      { S7_GenerateENO := "TRUE" } Add(in1 := "Archiwizowane_parametry".Wilgotnosc_srednia[0], in2 := "Archiwizowane_parametry".Wilgotnosc["Archiwizowane_parametry".iterator_srednia], out => "Archiwizowane_parametry".Wilgotnosc_srednia[0])
      Div(in1 := "Archiwizowane_parametry".Naslonecznienie_suma[0], in2 := "Archiwizowane_parametry".dzielnik, out => "Archiwizowane_parametry".Naslonecznienie_srednia[0])
      Div(in1 := "Archiwizowane_parametry".Temperatura_suma[0], in2 := "Archiwizowane_parametry".dzielnik, out => "Archiwizowane_parametry".Temperatura_srednia[0])
      Div(in1 := "Archiwizowane_parametry".Wilgotnosc_suma[0], in2 := "Archiwizowane_parametry".dzielnik, out => "Archiwizowane_parametry".Wilgotnosc_srednia[0])
   END_RUNG
   RUNG wire#w2
      { S7_Templates := "SrcType := Int" } GE_Contact(in1 := "Archiwizowane_parametry".iterator_srednia, in2 := 16)
      { S7_Templates := "SrcType := Int" } LT_Contact(in1 := "Archiwizowane_parametry".iterator_srednia, in2 := 32)
      { S7_GenerateENO := "TRUE" } Add(in1 := "Archiwizowane_parametry".Naslonecznienie_srednia[1], in2 := "Archiwizowane_parametry".Naslonecznienie["Archiwizowane_parametry".iterator_srednia], out => "Archiwizowane_parametry".Naslonecznienie_srednia[1])
      { S7_GenerateENO := "TRUE" } Add(in1 := "Archiwizowane_parametry".Temperatura_srednia[1], in2 := "Archiwizowane_parametry".Temperatura["Archiwizowane_parametry".iterator_srednia], out => "Archiwizowane_parametry".Temperatura_srednia[1])
      { S7_GenerateENO := "TRUE" } Add(in1 := "Archiwizowane_parametry".Wilgotnosc_srednia[1], in2 := "Archiwizowane_parametry".Wilgotnosc["Archiwizowane_parametry".iterator_srednia], out => "Archiwizowane_parametry".Wilgotnosc_srednia[1])
      Div(in1 := "Archiwizowane_parametry".Naslonecznienie_suma[1], in2 := "Archiwizowane_parametry".dzielnik, out => "Archiwizowane_parametry".Naslonecznienie_srednia[1])
      Div(in1 := "Archiwizowane_parametry".Temperatura_suma[1], in2 := "Archiwizowane_parametry".dzielnik, out => "Archiwizowane_parametry".Temperatura_srednia[1])
      Div(in1 := "Archiwizowane_parametry".Wilgotnosc_suma[1], in2 := "Archiwizowane_parametry".dzielnik, out => "Archiwizowane_parametry".Wilgotnosc_srednia[1])
   END_RUNG
   RUNG wire#w2
      { S7_Templates := "SrcType := Int" } GE_Contact(in1 := "Archiwizowane_parametry".iterator_srednia, in2 := 32)
      { S7_Templates := "SrcType := Int" } LT_Contact(in1 := "Archiwizowane_parametry".iterator_srednia, in2 := 48)
      { S7_GenerateENO := "TRUE" } Add(in1 := "Archiwizowane_parametry".Naslonecznienie_srednia[2], in2 := "Archiwizowane_parametry".Naslonecznienie["Archiwizowane_parametry".iterator_srednia], out => "Archiwizowane_parametry".Naslonecznienie_srednia[2])
      { S7_GenerateENO := "TRUE" } Add(in1 := "Archiwizowane_parametry".Temperatura_srednia[2], in2 := "Archiwizowane_parametry".Temperatura["Archiwizowane_parametry".iterator_srednia], out => "Archiwizowane_parametry".Temperatura_srednia[2])
      { S7_GenerateENO := "TRUE" } Add(in1 := "Archiwizowane_parametry".Wilgotnosc_srednia[2], in2 := "Archiwizowane_parametry".Wilgotnosc["Archiwizowane_parametry".iterator_srednia], out => "Archiwizowane_parametry".Wilgotnosc_srednia[2])
      Div(in1 := "Archiwizowane_parametry".Naslonecznienie_suma[2], in2 := "Archiwizowane_parametry".dzielnik, out => "Archiwizowane_parametry".Naslonecznienie_srednia[2])
      Div(in1 := "Archiwizowane_parametry".Temperatura_suma[2], in2 := "Archiwizowane_parametry".dzielnik, out => "Archiwizowane_parametry".Temperatura_srednia[2])
      Div(in1 := "Archiwizowane_parametry".Wilgotnosc_suma[2], in2 := "Archiwizowane_parametry".dzielnik, out => "Archiwizowane_parametry".Wilgotnosc_srednia[2])
   END_RUNG
   RUNG wire#w2
      { S7_Templates := "SrcType := Int" } GE_Contact(in1 := "Archiwizowane_parametry".iterator_srednia, in2 := 48)
      { S7_Templates := "SrcType := Int" } LT_Contact(in1 := "Archiwizowane_parametry".iterator_srednia, in2 := 64)
      { S7_GenerateENO := "TRUE" } Add(in1 := "Archiwizowane_parametry".Naslonecznienie_srednia[3], in2 := "Archiwizowane_parametry".Naslonecznienie["Archiwizowane_parametry".iterator_srednia], out => "Archiwizowane_parametry".Naslonecznienie_srednia[3])
      { S7_GenerateENO := "TRUE" } Add(in1 := "Archiwizowane_parametry".Temperatura_srednia[3], in2 := "Archiwizowane_parametry".Temperatura["Archiwizowane_parametry".iterator_srednia], out => "Archiwizowane_parametry".Temperatura_srednia[3])
      { S7_GenerateENO := "TRUE" } Add(in1 := "Archiwizowane_parametry".Wilgotnosc_srednia[3], in2 := "Archiwizowane_parametry".Wilgotnosc["Archiwizowane_parametry".iterator_srednia], out => "Archiwizowane_parametry".Wilgotnosc_srednia[3])
      Div(in1 := "Archiwizowane_parametry".Naslonecznienie_suma[3], in2 := "Archiwizowane_parametry".dzielnik, out => "Archiwizowane_parametry".Naslonecznienie_srednia[3])
      Div(in1 := "Archiwizowane_parametry".Temperatura_suma[3], in2 := "Archiwizowane_parametry".dzielnik, out => "Archiwizowane_parametry".Temperatura_srednia[3])
      Div(in1 := "Archiwizowane_parametry".Wilgotnosc_suma[3], in2 := "Archiwizowane_parametry".dzielnik, out => "Archiwizowane_parametry".Wilgotnosc_srednia[3])
   END_RUNG
   RUNG wire#w2
      { S7_Templates := "SrcType := Int" } GE_Contact(in1 := "Archiwizowane_parametry".iterator_srednia, in2 := 64)
      { S7_Templates := "SrcType := Int" } LT_Contact(in1 := "Archiwizowane_parametry".iterator_srednia, in2 := 80)
      { S7_GenerateENO := "TRUE" } Add(in1 := "Archiwizowane_parametry".Naslonecznienie_srednia[4], in2 := "Archiwizowane_parametry".Naslonecznienie["Archiwizowane_parametry".iterator_srednia], out => "Archiwizowane_parametry".Naslonecznienie_srednia[4])
      { S7_GenerateENO := "TRUE" } Add(in1 := "Archiwizowane_parametry".Temperatura_srednia[4], in2 := "Archiwizowane_parametry".Temperatura["Archiwizowane_parametry".iterator_srednia], out => "Archiwizowane_parametry".Temperatura_srednia[4])
      { S7_GenerateENO := "TRUE" } Add(in1 := "Archiwizowane_parametry".Wilgotnosc_srednia[4], in2 := "Archiwizowane_parametry".Wilgotnosc["Archiwizowane_parametry".iterator_srednia], out => "Archiwizowane_parametry".Wilgotnosc_srednia[4])
      Div(in1 := "Archiwizowane_parametry".Naslonecznienie_suma[4], in2 := "Archiwizowane_parametry".dzielnik, out => "Archiwizowane_parametry".Naslonecznienie_srednia[4])
      Div(in1 := "Archiwizowane_parametry".Temperatura_suma[4], in2 := "Archiwizowane_parametry".dzielnik, out => "Archiwizowane_parametry".Temperatura_srednia[4])
      Div(in1 := "Archiwizowane_parametry".Wilgotnosc_suma[4], in2 := "Archiwizowane_parametry".dzielnik, out => "Archiwizowane_parametry".Wilgotnosc_srednia[4])
   END_RUNG
   RUNG wire#w2
      { S7_Templates := "SrcType := Int" } GE_Contact(in1 := "Archiwizowane_parametry".iterator_srednia, in2 := 80)
      { S7_Templates := "SrcType := Int" } LT_Contact(in1 := "Archiwizowane_parametry".iterator_srednia, in2 := 96)
      { S7_GenerateENO := "TRUE" } Add(in1 := "Archiwizowane_parametry".Naslonecznienie_srednia[5], in2 := "Archiwizowane_parametry".Naslonecznienie["Archiwizowane_parametry".iterator_srednia], out => "Archiwizowane_parametry".Naslonecznienie_srednia[5])
      { S7_GenerateENO := "TRUE" } Add(in1 := "Archiwizowane_parametry".Temperatura_srednia[5], in2 := "Archiwizowane_parametry".Temperatura["Archiwizowane_parametry".iterator_srednia], out => "Archiwizowane_parametry".Temperatura_srednia[5])
      { S7_GenerateENO := "TRUE" } Add(in1 := "Archiwizowane_parametry".Wilgotnosc_srednia[5], in2 := "Archiwizowane_parametry".Wilgotnosc["Archiwizowane_parametry".iterator_srednia], out => "Archiwizowane_parametry".Wilgotnosc_srednia[5])
      Div(in1 := "Archiwizowane_parametry".Naslonecznienie_suma[5], in2 := "Archiwizowane_parametry".dzielnik, out => "Archiwizowane_parametry".Naslonecznienie_srednia[5])
      Div(in1 := "Archiwizowane_parametry".Temperatura_suma[5], in2 := "Archiwizowane_parametry".dzielnik, out => "Archiwizowane_parametry".Temperatura_srednia[5])
      Div(in1 := "Archiwizowane_parametry".Wilgotnosc_suma[5], in2 := "Archiwizowane_parametry".dzielnik, out => "Archiwizowane_parametry".Wilgotnosc_srednia[5])
   END_RUNG
   RUNG wire#w2
      { S7_Templates := "SrcType := Int" } GE_Contact(in1 := "Archiwizowane_parametry".iterator_srednia, in2 := 96)
      { S7_GenerateENO := "TRUE" } Add(in1 := "Archiwizowane_parametry".Naslonecznienie_srednia[6], in2 := "Archiwizowane_parametry".Naslonecznienie["Archiwizowane_parametry".iterator_srednia], out => "Archiwizowane_parametry".Naslonecznienie_srednia[6])
      { S7_GenerateENO := "TRUE" } Add(in1 := "Archiwizowane_parametry".Temperatura_srednia[6], in2 := "Archiwizowane_parametry".Temperatura["Archiwizowane_parametry".iterator_srednia], out => "Archiwizowane_parametry".Temperatura_srednia[6])
      { S7_GenerateENO := "TRUE" } Add(in1 := "Archiwizowane_parametry".Wilgotnosc_srednia[6], in2 := "Archiwizowane_parametry".Wilgotnosc["Archiwizowane_parametry".iterator_srednia], out => "Archiwizowane_parametry".Wilgotnosc_srednia[6])
      Div(in1 := "Archiwizowane_parametry".Naslonecznienie_suma[6], in2 := "Archiwizowane_parametry".dzielnik, out => "Archiwizowane_parametry".Naslonecznienie_srednia[6])
      Div(in1 := "Archiwizowane_parametry".Temperatura_suma[6], in2 := "Archiwizowane_parametry".dzielnik, out => "Archiwizowane_parametry".Temperatura_srednia[6])
      Div(in1 := "Archiwizowane_parametry".Wilgotnosc_suma[6], in2 := "Archiwizowane_parametry".dzielnik, out => "Archiwizowane_parametry".Wilgotnosc_srednia[6])
   END_RUNG
   RUNG wire#w1
      { S7_GenerateENO := "TRUE" } Add(in1 := "Archiwizowane_parametry".iterator_srednia, in2 := 1, out => "Archiwizowane_parametry".iterator_srednia)
   END_RUNG
   // the same network as SCL:
   // ENO of a box is taken as its EN; it also drops when the box reports an error
   #_w1 := "Archiwizowane_parametry".iterator_srednia < 112;
   #_w2 := #_w1 AND ("Archiwizowane_parametry".Wilgotnosc["Archiwizowane_parametry".iterator_srednia] >= 0);
   IF #_w2 THEN "Archiwizowane_parametry".dzielnik := "Archiwizowane_parametry".dzielnik + 1; END_IF;
   IF #_w2 AND ("Archiwizowane_parametry".iterator_srednia < 16) THEN
       "Archiwizowane_parametry".Naslonecznienie_srednia[0] := "Archiwizowane_parametry".Naslonecznienie_srednia[0] + "Archiwizowane_parametry".Naslonecznienie["Archiwizowane_parametry".iterator_srednia];
       "Archiwizowane_parametry".Temperatura_srednia[0] := "Archiwizowane_parametry".Temperatura_srednia[0] + "Archiwizowane_parametry".Temperatura["Archiwizowane_parametry".iterator_srednia];
       "Archiwizowane_parametry".Wilgotnosc_srednia[0] := "Archiwizowane_parametry".Wilgotnosc_srednia[0] + "Archiwizowane_parametry".Wilgotnosc["Archiwizowane_parametry".iterator_srednia];
       "Archiwizowane_parametry".Naslonecznienie_srednia[0] := "Archiwizowane_parametry".Naslonecznienie_suma[0] / "Archiwizowane_parametry".dzielnik;
       "Archiwizowane_parametry".Temperatura_srednia[0] := "Archiwizowane_parametry".Temperatura_suma[0] / "Archiwizowane_parametry".dzielnik;
       "Archiwizowane_parametry".Wilgotnosc_srednia[0] := "Archiwizowane_parametry".Wilgotnosc_suma[0] / "Archiwizowane_parametry".dzielnik;
   END_IF;
   IF #_w2 AND ("Archiwizowane_parametry".iterator_srednia >= 16) AND ("Archiwizowane_parametry".iterator_srednia < 32) THEN
       "Archiwizowane_parametry".Naslonecznienie_srednia[1] := "Archiwizowane_parametry".Naslonecznienie_srednia[1] + "Archiwizowane_parametry".Naslonecznienie["Archiwizowane_parametry".iterator_srednia];
       "Archiwizowane_parametry".Temperatura_srednia[1] := "Archiwizowane_parametry".Temperatura_srednia[1] + "Archiwizowane_parametry".Temperatura["Archiwizowane_parametry".iterator_srednia];
       "Archiwizowane_parametry".Wilgotnosc_srednia[1] := "Archiwizowane_parametry".Wilgotnosc_srednia[1] + "Archiwizowane_parametry".Wilgotnosc["Archiwizowane_parametry".iterator_srednia];
       "Archiwizowane_parametry".Naslonecznienie_srednia[1] := "Archiwizowane_parametry".Naslonecznienie_suma[1] / "Archiwizowane_parametry".dzielnik;
       "Archiwizowane_parametry".Temperatura_srednia[1] := "Archiwizowane_parametry".Temperatura_suma[1] / "Archiwizowane_parametry".dzielnik;
       "Archiwizowane_parametry".Wilgotnosc_srednia[1] := "Archiwizowane_parametry".Wilgotnosc_suma[1] / "Archiwizowane_parametry".dzielnik;
   END_IF;
   IF #_w2 AND ("Archiwizowane_parametry".iterator_srednia >= 32) AND ("Archiwizowane_parametry".iterator_srednia < 48) THEN
       "Archiwizowane_parametry".Naslonecznienie_srednia[2] := "Archiwizowane_parametry".Naslonecznienie_srednia[2] + "Archiwizowane_parametry".Naslonecznienie["Archiwizowane_parametry".iterator_srednia];
       "Archiwizowane_parametry".Temperatura_srednia[2] := "Archiwizowane_parametry".Temperatura_srednia[2] + "Archiwizowane_parametry".Temperatura["Archiwizowane_parametry".iterator_srednia];
       "Archiwizowane_parametry".Wilgotnosc_srednia[2] := "Archiwizowane_parametry".Wilgotnosc_srednia[2] + "Archiwizowane_parametry".Wilgotnosc["Archiwizowane_parametry".iterator_srednia];
       "Archiwizowane_parametry".Naslonecznienie_srednia[2] := "Archiwizowane_parametry".Naslonecznienie_suma[2] / "Archiwizowane_parametry".dzielnik;
       "Archiwizowane_parametry".Temperatura_srednia[2] := "Archiwizowane_parametry".Temperatura_suma[2] / "Archiwizowane_parametry".dzielnik;
       "Archiwizowane_parametry".Wilgotnosc_srednia[2] := "Archiwizowane_parametry".Wilgotnosc_suma[2] / "Archiwizowane_parametry".dzielnik;
   END_IF;
   IF #_w2 AND ("Archiwizowane_parametry".iterator_srednia >= 48) AND ("Archiwizowane_parametry".iterator_srednia < 64) THEN
       "Archiwizowane_parametry".Naslonecznienie_srednia[3] := "Archiwizowane_parametry".Naslonecznienie_srednia[3] + "Archiwizowane_parametry".Naslonecznienie["Archiwizowane_parametry".iterator_srednia];
       "Archiwizowane_parametry".Temperatura_srednia[3] := "Archiwizowane_parametry".Temperatura_srednia[3] + "Archiwizowane_parametry".Temperatura["Archiwizowane_parametry".iterator_srednia];
       "Archiwizowane_parametry".Wilgotnosc_srednia[3] := "Archiwizowane_parametry".Wilgotnosc_srednia[3] + "Archiwizowane_parametry".Wilgotnosc["Archiwizowane_parametry".iterator_srednia];
       "Archiwizowane_parametry".Naslonecznienie_srednia[3] := "Archiwizowane_parametry".Naslonecznienie_suma[3] / "Archiwizowane_parametry".dzielnik;
       "Archiwizowane_parametry".Temperatura_srednia[3] := "Archiwizowane_parametry".Temperatura_suma[3] / "Archiwizowane_parametry".dzielnik;
       "Archiwizowane_parametry".Wilgotnosc_srednia[3] := "Archiwizowane_parametry".Wilgotnosc_suma[3] / "Archiwizowane_parametry".dzielnik;
   END_IF;
   IF #_w2 AND ("Archiwizowane_parametry".iterator_srednia >= 64) AND ("Archiwizowane_parametry".iterator_srednia < 80) THEN
       "Archiwizowane_parametry".Naslonecznienie_srednia[4] := "Archiwizowane_parametry".Naslonecznienie_srednia[4] + "Archiwizowane_parametry".Naslonecznienie["Archiwizowane_parametry".iterator_srednia];
       "Archiwizowane_parametry".Temperatura_srednia[4] := "Archiwizowane_parametry".Temperatura_srednia[4] + "Archiwizowane_parametry".Temperatura["Archiwizowane_parametry".iterator_srednia];
       "Archiwizowane_parametry".Wilgotnosc_srednia[4] := "Archiwizowane_parametry".Wilgotnosc_srednia[4] + "Archiwizowane_parametry".Wilgotnosc["Archiwizowane_parametry".iterator_srednia];
       "Archiwizowane_parametry".Naslonecznienie_srednia[4] := "Archiwizowane_parametry".Naslonecznienie_suma[4] / "Archiwizowane_parametry".dzielnik;
       "Archiwizowane_parametry".Temperatura_srednia[4] := "Archiwizowane_parametry".Temperatura_suma[4] / "Archiwizowane_parametry".dzielnik;
       "Archiwizowane_parametry".Wilgotnosc_srednia[4] := "Archiwizowane_parametry".Wilgotnosc_suma[4] / "Archiwizowane_parametry".dzielnik;
   END_IF;
   IF #_w2 AND ("Archiwizowane_parametry".iterator_srednia >= 80) AND ("Archiwizowane_parametry".iterator_srednia < 96) THEN
       "Archiwizowane_parametry".Naslonecznienie_srednia[5] := "Archiwizowane_parametry".Naslonecznienie_srednia[5] + "Archiwizowane_parametry".Naslonecznienie["Archiwizowane_parametry".iterator_srednia];
       "Archiwizowane_parametry".Temperatura_srednia[5] := "Archiwizowane_parametry".Temperatura_srednia[5] + "Archiwizowane_parametry".Temperatura["Archiwizowane_parametry".iterator_srednia];
       "Archiwizowane_parametry".Wilgotnosc_srednia[5] := "Archiwizowane_parametry".Wilgotnosc_srednia[5] + "Archiwizowane_parametry".Wilgotnosc["Archiwizowane_parametry".iterator_srednia];
       "Archiwizowane_parametry".Naslonecznienie_srednia[5] := "Archiwizowane_parametry".Naslonecznienie_suma[5] / "Archiwizowane_parametry".dzielnik;
       "Archiwizowane_parametry".Temperatura_srednia[5] := "Archiwizowane_parametry".Temperatura_suma[5] / "Archiwizowane_parametry".dzielnik;
       "Archiwizowane_parametry".Wilgotnosc_srednia[5] := "Archiwizowane_parametry".Wilgotnosc_suma[5] / "Archiwizowane_parametry".dzielnik;
   END_IF;
   IF #_w2 AND ("Archiwizowane_parametry".iterator_srednia >= 96) THEN
       "Archiwizowane_parametry".Naslonecznienie_srednia[6] := "Archiwizowane_parametry".Naslonecznienie_srednia[6] + "Archiwizowane_parametry".Naslonecznienie["Archiwizowane_parametry".iterator_srednia];
       "Archiwizowane_parametry".Temperatura_srednia[6] := "Archiwizowane_parametry".Temperatura_srednia[6] + "Archiwizowane_parametry".Temperatura["Archiwizowane_parametry".iterator_srednia];
       "Archiwizowane_parametry".Wilgotnosc_srednia[6] := "Archiwizowane_parametry".Wilgotnosc_srednia[6] + "Archiwizowane_parametry".Wilgotnosc["Archiwizowane_parametry".iterator_srednia];
       "Archiwizowane_parametry".Naslonecznienie_srednia[6] := "Archiwizowane_parametry".Naslonecznienie_suma[6] / "Archiwizowane_parametry".dzielnik;
       "Archiwizowane_parametry".Temperatura_srednia[6] := "Archiwizowane_parametry".Temperatura_suma[6] / "Archiwizowane_parametry".dzielnik;
       "Archiwizowane_parametry".Wilgotnosc_srednia[6] := "Archiwizowane_parametry".Wilgotnosc_suma[6] / "Archiwizowane_parametry".dzielnik;
   END_IF;
   IF #_w1 THEN
       "Archiwizowane_parametry".iterator_srednia := "Archiwizowane_parametry".iterator_srednia + 1;
   END_IF;
END_REGION
END_FUNCTION

// folder: LGF/4 Math operations

FUNCTION "LGF_RandomRange_Real" : Real   // FC10014, SCL
TITLE = LGF_RandomRange_Real
{ S7_Optimized_Access := 'TRUE' }
AUTHOR : Siemens_Digital_Industries
FAMILY : LGF
NAME : LGF_RandomRange_Real
// This function generates random numbers in defined limits (Datatype Real)
   VAR_INPUT
      minValue : Real;   // minimal Value random can reach / Minimum value of the range of the random number
      maxValue : Real;   // maximal Value random can reach / Maximum value of the range of the random number
   END_VAR
   VAR_OUTPUT
      error : Bool;   // Error if true
      status : Word;   // Status of the function
      subfunctionStatus : Word;   // Status or return value of called FB's, FCs and system blocks
   END_VAR
   VAR_TEMP
      tempTime : DTL;   // System time
      tempNanoSecondInDWord : DWord;   // UDINT converted to DWORD for access to individual bytes
      tempTimeStatus : Word;   // Status of the instruction RD_SYS_T
      tempRandomValue : DWord;   // Random-start-value
      tempNormReal : Real;   // normalized value
   END_VAR
   // Ret_Val : Returns random Real number in predefined range
   VAR CONSTANT
      ZERO : Real := 0.0;   // Zero value in case of error
      MAX_UDINT : UDInt := 4294967295;   // Maximum UDINT value
      SUB_STATUS_NO_ERROR : Word := 16#0000;   // Status: sub function call ends without error
      STATUS_FINISHED_NO_ERROR : Word := 16#0000;   // Status: Execution finished without errors
      ERR_MAX_LESS_MIN : Word := 16#8200;   // Error: The maximum limit number is smaller than the minimum limit number
      ERR_RD_SYS_T : Word := 16#8600;   // Error: System function Read system time returned an error
   END_VAR
BEGIN
   REGION Block info header
     //=============================================================================
     // SIEMENS AG / (c)Copyright 2017
     //-----------------------------------------------------------------------------
     // Title:            LGF_RandomRange_Real
     // Comment/Function: This function generates random numbers in defined limits (Datatype Real)
     // Library/Family:   LGF(Library General Functions)
     // Author:           Siemens Digital Industry Support
     // Tested with:      S7-PLCSIM Advanced V2.0 SP1
     // Engineering:      TIA Portal V15 Update 2
     // Restrictions:     ENO disabled - error handling done by error and status
     // Requirements:     PLC (S7-1200 / S7-1500)
     //-------------------------------------------------------------------------------
     // Change log table:
     // Version  | Date       | Expert in charge       | Changes applied
     //----------|------------|------------------------|------------------------------
     // 01.00.00 19.08.2015  Siemens Industry Online Support
     //                      First released version
     // 01.00.01 02.01.2017  Siemens Industry Online Support
     //                      Upgrade: TIA Portal V14 Update 1
     // 01.00.02 02.03.2017  Siemens Industry Online Support
     //                      Bugfix: FC number
     // 01.00.03 17.08.2018  Siemens Industry Online Support
     //                      Upgrade: TIA V15 Update 2
     // 01.00.04 23.11.2018  Siemens Industry Online Support
     //                      Upgrade: TIA V15.1
     // 01.01.00 13.11.2019  Siemens Industry Presales Support
     //                      Renamed from "LGF_RandomReal" to "LGF_RandomRange_Real"
     //                      Regions, commens and costants are added
     // 03.00.00 23.04.2020  Siemens Industry Support
     //                      Set version to V3.0.0, harmonize the version of the whole library
     //=============================================================================
   END_REGION

   REGION Validation
     // Check if the maximal Value is less than the minimal value
     IF (#minValue > #maxValue) THEN
       #error := true;
       #status := #ERR_MAX_LESS_MIN;
       #subfunctionStatus := #SUB_STATUS_NO_ERROR;
       #LGF_RandomRange_Real := #ZERO;
       RETURN;
     END_IF;

     // Read system time
     #tempTimeStatus := INT_TO_WORD(RD_SYS_T(#tempTime));

     // Check return variable for error
     IF (#tempTimeStatus <> #SUB_STATUS_NO_ERROR) THEN
       #error := true;
       #status := #ERR_RD_SYS_T;
       #subfunctionStatus := #tempTimeStatus;
       #LGF_RandomRange_Real := #ZERO;
       RETURN;
     END_IF;
   END_REGION

   REGION Calculating random number
     // Converting to double word so individual bytes can be addressed
     #tempNanoSecondInDWord := UDINT_TO_DWORD(#tempTime.NANOSECOND);

     // Calculate a random-start-value depending on the time
     #tempRandomValue.%B3 := #tempNanoSecondInDWord.%B0;
     #tempRandomValue.%B2 := #tempNanoSecondInDWord.%B1;
     #tempRandomValue.%B1 := #tempNanoSecondInDWord.%B2;
     #tempRandomValue.%B0 := #tempNanoSecondInDWord.%B3;

     // Norm the calculated random number: 0.0 <= #tempNormReal <= 1.0
     #tempNormReal := UDINT_TO_REAL(DWORD_TO_UDINT(#tempRandomValue)) / UDINT_TO_REAL(#MAX_UDINT);

     // Scale the tempNormReal to be in the range of maxValue and minValue
     #LGF_RandomRange_Real := ((#tempNormReal * (#maxValue - #minValue) + (#minValue)));

     #error := false;
     #status := #STATUS_FINISHED_NO_ERROR;
     #subfunctionStatus := #SUB_STATUS_NO_ERROR;
     // ENO mechanism is not used
     ENO := TRUE;
   END_REGION
END_FUNCTION

// ===== PLC "PLC_Web_server"  CPU 1518-4 PN/DP =====

VAR_GLOBAL   // PLC tag table "Default tag table"
   "err" AT %MW1 : Int;
   "tag1" AT %M6.0 : Bool;
END_VAR

DATA_BLOCK "Wejscia_PLC"   // DB2
{ S7_Optimized_Access := 'TRUE' }
VERSION : 0.1
   VAR
      Czujnik_wilgotności_powietrza : Int;   // Czujnik wilgotności powietrza w szklarni
      Czujnik_wilgotności_gleby : Int;   // Czujnik wilgotności gleby w szklarni
      Temperatura_wewnetrzna : Real;   // Temperatura wewnątrz szklarni
      Czujnik_natezenia_swiatła : Int;   // Czujnik natężenia światła wewnątrz szklarni
      Wewnetrzny_czujnik_CO2 : Int;   // Czujnik stężenia dwutlenku węgla w szklarni
      Stopien_zasloniecia_rolet : Int;   // Stopień zasłonięcia rolet w szklarni (przyjęty przedział 0-100%)
   END_VAR
BEGIN
END_DATA_BLOCK

// folder: Archiwizacja_parametrow

DATA_BLOCK "Archiwizowane_parametry"   // DB4
{ S7_Optimized_Access := 'TRUE' }
VERSION : 0.1
   VAR
      Temperatura : Array[0..111] of Real;
      Wilgotnosc : Array[0..111] of Int;
      Naslonecznienie : Array[0..111] of Int;
      iterator : Int := 0;   // Iterator służący do zapisu danych w odpowiednich komórkach tablicy.
   END_VAR
BEGIN
   Naslonecznienie[0] := 0;
   Naslonecznienie[1] := 0;
END_DATA_BLOCK

// folder: (top level)

ORGANIZATION_BLOCK "Main"   // OB1, LAD, ProgramCycle
TITLE = "Main Program Sweep (Cycle)"
{ S7_Optimized_Access := 'TRUE' }
VERSION : 0.1
   VAR_INPUT
      Initial_Call : Bool;   // Initial call of this OB
      Remanence : Bool;   // =True, if remanent data are available
   END_VAR
BEGIN

REGION Network 1
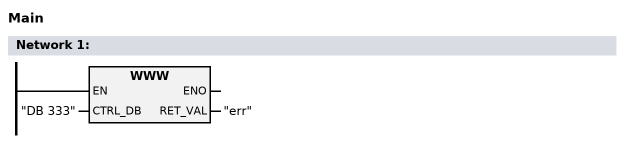
   "err" := WWW(CTRL_DB := "DB 333");
END_REGION
END_ORGANIZATION_BLOCK

(* ===== HMI "HMI_RT_3" =====
system functions are stored by id; their names below are inferred from use
connection "HMI_Connection_4": ETHERNET, SMART_S7_1200_OMS

HMI tags "Default tag table"
   "AlwaysTRUE" : Bool = PLC AlwaysTRUE AT %M1.2, 1 s
   "Grzałka" : Bool = PLC Grzałka AT %Q0.0, 1 s
   "HMI_Aktywacja_trybu_automatycznego" : Bool = PLC HMI.Aktywacja_trybu_automatycznego, 1 s
   "HMI_Aktywacja_trybu_Receptur" : Bool = PLC HMI.Aktywacja_trybu_Receptur, 1 s
   "HMI_Aktywacja_trybu_zapis_Receptur" : Bool = PLC HMI.Aktywacja_trybu_zapis_Receptur, 1 s
   "HMI_Reset_Trybow" : Bool = PLC HMI.Reset_Trybow, 1 s
   "Pompa_podlewanie" : Bool = PLC Pompa_podlewanie AT %Q1.0, 1 s
   "Pompa_zraszacze" : Bool = PLC Pompa_zraszacze AT %Q0.2, 1 s
   "Tag_ScreenNumber" : Int = PLC HMI.Numer_ekranu_HMI AT %MD0, 100 ms
   "Tryb_auto_parametry_Naslonecznienie" : Int = PLC Tryb_auto_parametry.Naslonecznienie, 1 s
   "Tryb_auto_parametry_Stezenie_co2" : Int = PLC Tryb_auto_parametry.Stezenie_co2, 1 s
   "Tryb_auto_parametry_System_okien" : Bool = PLC Tryb_auto_parametry.System_okien, 1 s
   "Tryb_auto_parametry_Temperatura" : Real = PLC Tryb_auto_parametry.Temperatura, 1 s
   "Tryb_auto_parametry_Wilgotnosc_gleby" : Int = PLC Tryb_auto_parametry.Wilgotnosc_gleby, 1 s
   "Tryb_auto_parametry_Wilgotnosc_powietrza" : Int = PLC Tryb_auto_parametry.Wilgotnosc_powietrza, 1 s
   "Wentylator" : Bool = PLC Wentylator AT %Q0.1, 1 s

HMI tags "Z_PLC"
   "Czujnik_wilgotności_powietrza" : Int = PLC Wejscia_PLC.Czujnik_wilgotności_powietrza, 500 ms
   "Temperatura_wewnetrzna" : Real = PLC Wejscia_PLC.Temperatura_wewnetrzna, 500 ms
   "Czujnik_natezenia_światła" : Int = PLC Wejscia_PLC.Czujnik_natezenia_swiatła, 500 ms
   "Czujnik_wilgotności_gleby" : Int = PLC Wejscia_PLC.Czujnik_wilgotności_gleby, 500 ms
   "Wewnetrzny_czujnik_CO2" : Int = PLC Wejscia_PLC.Wewnetrzny_czujnik_CO2, 500 ms
   "Czujnik_wiatru" : Int = PLC Wejscia_PLC.Czujnik_wiatru, 500 ms
   "Stopien_zasloniecia_rolet" : Int = PLC Wejscia_PLC.Stopien_zasloniecia_rolet, 1 s
   "Zewnetrzny_czujnik_CO2" : Int = PLC Wejscia_PLC.Zewnetrzny_czujnik_CO2 AT %DB1.DBW0, 1 s
   "Temperatura_zewnetrzna" : Real = PLC Wejscia_PLC.Temperatura_zewnetrzna AT %DB1.DBW0, 1 s

HMI tags "Do_PLC"
   "System_okien_auto" : Bool = PLC HMI.System_okien_auto, 500 ms
   "Stopien_zasloniecia_rolet_manual" : Int = PLC HMI.Stopien_zasloniecia_rolet_manual, 100 ms
   "Przycisk_zraszania_manual" : Bool = PLC HMI.Przycisk_zraszacze_manual AT %Q0.2, 100 ms
   "Przycisk_wentylacja_manual" : Bool = PLC HMI.Przycisk_wentylacja_manual AT %Q0.1, 100 ms
   "Przycisk_grzanie_manual" : Bool = PLC HMI.Przycisk_grzanie_manual AT %Q0.0, 100 ms
   "Otwarcie_okien_man" : Bool = PLC HMI.Otwarcie_okien_manual AT %DB1.DBW0, 100 ms
   "Temperatura_auto" : Real = PLC HMI.Temperatura_auto, 500 ms
   "Naslonecznienie_auto" : Int = PLC HMI.Naslonecznienie_auto AT %DB1.DBW0, 500 ms
   "Wilgotnosc_powietrza_auto" : Int = PLC HMI.Wilgotnosc_powietrza_auto AT %DB1.DBW0, 500 ms
   "Wilgotnosc_gleby_auto" : Int = PLC HMI.Wilgotnosc_gleby_auto AT %DB1.DBW0, 500 ms
   "Przycisk_zatwierdz_auto" : Bool = PLC HMI.Przycisk_zatwierdz_auto AT %DB1.DBW0, 100 ms
   "nazwa_receptury" : String[254] = PLC HMI.nazwa_receptury AT %DB1.DBX0.0, 500 ms
   "przycisk_zatwierdz_zapis_receptury" : Bool = PLC HMI.Przycisk_zatwierdz_zapis_receptury AT %DB1.DBX0.0, 500 ms
   "HMI_Przycisk_zatwierdz_wybor_receptury" : Bool = PLC HMI.Przycisk_zatwierdz_wybor_receptury AT %DB1.DBX0.0, 500 ms
   "Przycisk_podlewania_manual" : Bool = PLC HMI.Przycisk_podlewanie_manual AT %Q0.2, 100 ms
   "Poziom_CO2_auto" : Int = PLC HMI.Poziom_CO2_auto AT %DB1.DBX0.0, 1 s

analog alarms
   3: 'Podmuchy wiatru osiągają wartości powyżej 35 km/h, system automatyczny zamyka okna.', class Warnings, trigger "Czujnik_wiatru"
   2: 'Temperatura powyżej 35 stopni / Temperatura powyżej 35 stopni, zaleca się wyłączenie grzania.', class Warnings, trigger "Temperatura_wewnetrzna"
   5: 'Temperatura powyżej 45 stopni, NIEZWŁOCZNIE SPRAWDŹ DZIAŁANIE GRZAŁKI, TERMOMETRU LUB WENTYLATORA. / Temperatura powyżej 45 stopni, NIEZWŁOCZNIE SPRAWDŹ DZIAŁANIE GRZAŁKI, TERMOMETRU LUB WENTYLATORA. JEŚLI TEMPERATURA NIE SPADA ZALECA SIĘ EWAKUOWAĆ WSZYSTKICH PRZEBYWAJĄCYCH W POMIESZCZENIU', class Errors, trigger "Temperatura_wewnetrzna"
   4: 'Stężenie CO2 ma powyżej 5000 jednostek. NIEZWŁOCZNIE OTWORZ OKNA ORAZ ZAŁĄCZ WENTYLATOR, NASTĘPNIE NALEŻY EWAKUOWAĆ WSZYSTKUCH ZNAJDUJĄCYCH SIĘ W POMIESZCZENIU / Stężenie CO2 ma powyżej 5000 jednostek. NIEZWŁOCZNIE OTWORZ OKNA ORAZ ZAŁĄCZ WENTYLATOR, NASTĘPNIE NALEŻY EWAKUOWAĆ WSZYSTKUCH ZNAJDUJĄCYCH SIĘ W POMIESZCZENIU', class Errors, trigger "Wewnetrzny_czujnik_CO2"
   1: 'Stężenie CO2 ma powyżej 3000 jednostek / Stężenie CO2 ma powyżej 3000 jednostek, dłużesze przebywanie w takim środowisku może być szkodliwe dla człowieka. Zalecane jest włączenie wentylacji lub otworzenie okien.', class Warnings, trigger "Wewnetrzny_czujnik_CO2"

text list "receptury": 0..1 ''

recipe "Receptura_nr1": Temperatura <- "Tryb_auto_parametry_Temperatura", Wilgotność Powietrza <- "Tryb_auto_parametry_Wilgotnosc_powietrza", Wilgotność gleby <- "Tryb_auto_parametry_Wilgotnosc_gleby", System okien <- "Tryb_auto_parametry_System_okien", Stężenie CO2 <- "Tryb_auto_parametry_Stezenie_co2", Nasłonecznienie <- "Tryb_auto_parametry_Naslonecznienie"

screen "tryb_manualny" 800x480
   on GenerateScreen: SetTag("Tag_ScreenNumber", 2)
   TextField "Text field_1" at 295,7 size 223x34; Text 'TRYB MANUALNY'
   TextField "Text field_4" at 512,155 size 171x61; Text 'STOPIEŃ OTWARCIA OKIEN OTWIERANIE OKIEN'
   Button "Button_4" at 518,261 size 80x70; TextOff 'PODLEWANIE'
      on Click: InvertBit("Przycisk_podlewania_manual")
   Button "Button_5" at 611,261 size 80x70; TextOff 'GRZANIE'
      on Click: InvertBit("Przycisk_grzanie_manual")
   Button "Button_6" at 701,261 size 80x70; TextOff 'WENTYLACJA'
      on Click: InvertBit("Przycisk_wentylacja_manual")
   GraphicView "Graphic view_1" at 710,356 size 60x60; Picture "fan_4829316"
      Visibility <- "Wentylator"
   GraphicView "Graphic view_6" at 622,356 size 60x60; Picture "heater_4463010"
      Visibility <- "Grzałka"
   GraphicView "Graphic view_7" at 527,356 size 64x60; Picture "irrigation_18631825"
      Visibility <- "Pompa_podlewanie"
   GraphicView "Graphic view_9" at 710,356 size 60x60; Picture "fan_off"
      Visibility <- "Wentylator"
   GraphicView "Graphic view_10" at 622,356 size 60x60; Picture "heater_off"
      Visibility <- "Grzałka"
   GraphicView "Graphic view_11" at 527,356 size 64x60; Picture "irrigation_off"
      Visibility <- "Pompa_podlewanie"
   Button "Button_14" at 6,7 size 43x43; TextOff 'DOM'; PictureOff "home_1"
      on Click: ActivateScreen("Root screen", 0)
   Button "Button_1" at 740,0 size 60x60; TextOff 'Text'; PictureOff "Back_arrow"
      on Click: function_efd93a16()
   Circle "Circle_1" at 541,428 size 42x42
      Visibility <- "Pompa_podlewanie"
   Circle "Circle_4" at 541,428 size 42x42
      Visibility <- "Pompa_podlewanie"
   Circle "Circle_2" at 631,428 size 42x42
      Visibility <- "Grzałka"
   Circle "Circle_5" at 631,428 size 42x42
      Visibility <- "Grzałka"
   Circle "Circle_3" at 720,428 size 41x41
      Visibility <- "Wentylator"
   Circle "Circle_6" at 720,428 size 41x41
      Visibility <- "Wentylator"
   TextField "Text field_8" at 405,71 size 117x61; Text 'STOPIEŃ OTWARCIA OKIEN STOPIEŃ ZASŁONIECIA ROLET'
   Bar "Bar_6" at 624,82 size 165x66; MinimumValue 0; MaximumValue 100
      ProcessValue <- "Stopien_zasloniecia_rolet_manual"
   Button "Button_3" at 530,114 size 80x50; TextOff '+ / ODSŁOŃ'
      on Click: function_b9b71300("Stopien_zasloniecia_rolet_manual", 5)
   Button "Button_7" at 530,60 size 80x50; TextOff '- / ZASŁOŃ'
      on Press: function_dd21b452("Stopien_zasloniecia_rolet_manual", 5)
   Button "Button_2" at 425,261 size 80x70; TextOff 'PODLEWANIE / MIKROZRASZANIE'
      on Click: InvertBit("Przycisk_zraszania_manual")
   GraphicView "Graphic view_2" at 434,356 size 60x60; Picture "sprinkler_4552152"
      Visibility <- "Pompa_zraszacze"
   GraphicView "Graphic view_3" at 434,356 size 60x60; Picture "sprinkler"
      Visibility <- "Pompa_zraszacze"
   Circle "Circle_7" at 443,428 size 42x42
      Visibility <- "Pompa_zraszacze"
   Circle "Circle_8" at 443,428 size 42x42
      Visibility <- "Pompa_zraszacze"
   Switch "Switch_1" at 499,199 size 209x37; TextOn 'OTWARTE'; CaptionText 'Switch'; TextOff 'ZAMKNIĘTE'
      ProcessValue <- "Otwarcie_okien_man"
   TextField "Text field_3" at 11,375 size 166x23; Text 'SZYBKOŚĆ WIATRU'
   IOField "I/O field_3" at 62,407 size 70x65; FormatPattern 999
      ProcessValue <- "Czujnik_wiatru"
   IOField "I/O field_1" at 48,189 size 101x32; FormatPattern 99999
      ProcessValue <- "Czujnik_natezenia_światła"
   TextField "Text field_15" at 129,408 size 52x72; Text 'Km h'
   IOField "I/O field_2" at 44,292 size 83x65; FormatPattern 9999
      ProcessValue <- "Wewnetrzny_czujnik_CO2"
   TextField "Text field_11" at 118,301 size 69x39; Text 'ppm'
   TextField "Text field_5" at 14,148 size 204x23; Text 'INSOLATION / NASŁONECZNIENIE / SONNENEINSTRAHLUNG'
   IOField "I/O field_8" at 58,95 size 93x40; FormatPattern 99.99
      ProcessValue <- "Temperatura_wewnetrzna"
   TextField "Text field_20" at 30,56 size 137x42; Text 'TEMPERATURA TEMPERATURA WEWNTĘTRZNA'
   TextField "Text field_7" at 200,375 size 175x23; Text 'WILGOTNOŚĆ GLEBY'
   IOField "I/O field_5" at 248,293 size 83x65; FormatPattern 9999
      ProcessValue <- "Zewnetrzny_czujnik_CO2"
   IOField "I/O field_4" at 266,174 size 69x65; FormatPattern 999
      ProcessValue <- "Czujnik_wilgotności_powietrza"
   IOField "I/O field_6" at 261,405 size 68x65; FormatPattern 999
      ProcessValue <- "Czujnik_wilgotności_gleby"
   TextField "Text field_12" at 324,182 size 47x46; Text '%'
   TextField "Text field_13" at 321,416 size 47x46; Text '%'
   TextField "Text field_16" at 326,292 size 69x39; Text 'ppm'
   IOField "I/O field_9" at 248,85 size 97x65; FormatPattern 99.99
      ProcessValue <- "Temperatura_zewnetrzna"
   TextField "Text field_23" at 333,90 size 46x46; Text '°C'
   TextField "Text field_22" at 229,57 size 132x42; Text 'TEMPERATURA TEMPERATURA ZEWNĘTRZNA'
   TextField "Text field_9" at 229,256 size 123x42; Text 'STĘŻENIE CO2 ZEWNĘTRZNE STĘŻENIE CO2'
   TextField "Text field_6" at 180,143 size 223x42; Text 'WILGOTNOŚĆ POWIETRZA WILGOTNOŚĆ POWIETRZA'
   TextField "Text field_14" at 140,170 size 47x72; Text 'W m²'
   TextField "Text field_21" at 141,90 size 46x46; Text '°C'
   GraphicView "Graphic view_4" at 419,176 size 60x60; Picture "window_11250237"
   GraphicView "Graphic view_5" at 197,182 size 50x50; Picture "sensor_4212519"
   GraphicView "Graphic view_8" at 4,182 size 50x50; Picture "sensor_4212513"
   GraphicView "Graphic view_12" at 3,87 size 50x50; Picture "Thermometer_icon"
   GraphicView "Graphic view_13" at 199,87 size 50x50; Picture "Thermometer_icon"
   GraphicView "Graphic view_14" at 3,302 size 40x40; Picture "sensor_2828470"
   GraphicView "Graphic view_15" at 197,300 size 40x40; Picture "sensor_2828470"
   GraphicView "Graphic view_16" at 198,412 size 50x50; Picture "soil-sensor_11298794"
   GraphicView "Graphic view_17" at 3,416 size 50x50; Picture "anemometer_1113716"
   TextField "Text field_2" at 27,256 size 124x42; Text 'STĘŻENIE CO2 WEWNĘTRZNE STĘŻENIE CO2'

screen "tryb_automatyczny" 800x480
   on GenerateScreen: SetTag("Tag_ScreenNumber", 1)
   IOField "I/O field_1" at 67,322 size 57x40; FormatPattern 99.9
      ProcessValue <- "Temperatura_wewnetrzna"
   Button "Button_1" at 745,0 size 55x55; TextOff 'WRÓĆ'; PictureOff "Back_arrow"
      on Click: function_efd93a16()
   Button "Button_2" at 373,382 size 416x89; TextOff 'ZATWIERDŹ'
      on Click: ResetBit("HMI_Reset_Trybow"); SetBit("HMI_Aktywacja_trybu_automatycznego"); ActivateScreen("praca", 0)
   Bar "Bar_1" at 7,110 size 50x250; MinimumValue 0; MaximumValue 45
      ProcessValue <- "Temperatura_auto"
   TextField "Text field_2" at 1,71 size 132x23; Text 'TEMPERATURA'
   Bar "Bar_2" at 170,111 size 50x250; MinimumValue 0; MaximumValue 100
      ProcessValue <- "Wilgotnosc_powietrza_auto"
   TextField "Text field_3" at 165,68 size 122x42; Text 'WOLGOTNOŚĆ POWIETRZA WILGOTNOŚĆ POWIETRZA'
   Button "Button_3" at 71,115 size 75x45; TextOff '+ / +0.5 °C'
      on Press: function_dd21b452("Temperatura_auto", 0.5)
   Button "Button_7" at 71,183 size 75x45; TextOff '- / -0.5 °C'
      on Press: function_b9b71300("Temperatura_auto", 0.5)
   IOField "I/O field_2" at 67,251 size 62x40; FormatPattern 99.9
      ProcessValue <- "Temperatura_auto"
   TextField "Text field_11" at 122,260 size 23x22; Text '°C'
   TextField "Text field_9" at 122,333 size 23x22; Text '°C'
   Bar "Bar_4" at 335,111 size 50x250; MinimumValue 0; MaximumValue 100
      ProcessValue <- "Wilgotnosc_gleby_auto"
   TextField "Text field_10" at 332,65 size 122x42; Text 'WOLGOTNOŚĆ GLEBY WILGOTNOŚĆ GLEBY'
   Button "Button_8" at 398,132 size 65x40; TextOff '+ / +2%'
      on Click: function_dd21b452("Wilgotnosc_gleby_auto", 2)
   Button "Button_9" at 398,181 size 65x40; TextOff '- / -2%'
      on Click: function_b9b71300("Wilgotnosc_gleby_auto", 2)
   IOField "I/O field_5" at 402,255 size 60x40; FormatPattern 999
      ProcessValue <- "Wilgotnosc_gleby_auto"
   IOField "I/O field_6" at 404,325 size 58x40; FormatPattern 999
      ProcessValue <- "Czujnik_wilgotności_gleby"
   TextField "Text field_12" at 385,243 size 101x22; Text 'USTAWIONA'
   TextField "Text field_13" at 389,314 size 86x22; Text 'AKTUALNA'
   TextField "Text field_14" at 439,264 size 23x22; Text '%'
   TextField "Text field_15" at 439,335 size 23x22; Text '%'
   Button "Button_10" at 229,126 size 65x40; TextOff '+ / +5%'
      on Click: function_dd21b452("Wilgotnosc_powietrza_auto", 5)
   Button "Button_11" at 229,186 size 65x40; TextOff '- / -5%'
      on Click: function_b9b71300("Wilgotnosc_powietrza_auto", 5)
   IOField "I/O field_4" at 234,248 size 66x40; FormatPattern 999
      ProcessValue <- "Wilgotnosc_powietrza_auto"
   IOField "I/O field_7" at 236,320 size 62x40; FormatPattern 999
      ProcessValue <- "Czujnik_wilgotności_powietrza"
   TextField "Text field_16" at 223,235 size 101x22; Text 'USTAWIONA'
   TextField "Text field_17" at 223,306 size 86x22; Text 'AKTUALNA'
   TextField "Text field_18" at 275,257 size 23x22; Text '%'
   TextField "Text field_19" at 275,328 size 23x22; Text '%'
   Button "Button_14" at 4,7 size 45x45; TextOff 'DOM'; PictureOff "home_1"
      on Click: ActivateScreen("Root screen", 0)
   TextField "Text field_4" at 143,381 size 128x23; Text 'SYSTEM OKIEN'
   Switch "Switch_1" at 106,410 size 216x46; TextOn 'ON'; CaptionText 'Switch'; TextOff 'OFF'
      ProcessValue <- "System_okien_auto"
   GraphicView "Graphic view_1" at 129,70 size 40x40; Picture "Thermometer_icon"
   GraphicView "Graphic view_2" at 281,68 size 40x40; Picture "sensor_4212519"
   TextField "Text field_5" at 60,309 size 86x22; Text 'AKTUALNA'
   TextField "Text field_6" at 57,237 size 101x22; Text 'USTAWIONA'
   GraphicView "Graphic view_3" at 443,71 size 40x40; Picture "soil-sensor_11298794"
   TextField "Text field_1" at 255,4 size 291x47; Text 'TRYB AUTOMATYCZNY'
   Bar "Bar_3" at 496,111 size 50x250; MinimumValue 0; MaximumValue 1500
      ProcessValue <- "Naslonecznienie_auto"
   TextField "Text field_7" at 492,55 size 154x40; Text 'WOLGOTNOŚĆ GLEBY NASŁONECZNIENIE'
   GraphicView "Graphic view_4" at 585,86 size 40x40; Picture "sensor_4212513"
   Button "Button_4" at 553,131 size 82x43; TextOff '+ +50 W m'
      on Click: function_dd21b452("Naslonecznienie_auto", 50)
   Button "Button_5" at 554,186 size 82x43; TextOff '- -50 W m'
      on Click: function_b9b71300("Naslonecznienie_auto", 50)
   IOField "I/O field_3" at 561,254 size 61x40; FormatPattern 9999
      ProcessValue <- "Naslonecznienie_auto"
   TextField "Text field_8" at 545,242 size 101x22; Text 'USTAWIONA / USTAWIONE'
   IOField "I/O field_8" at 563,325 size 62x40; FormatPattern 9999
      ProcessValue <- "Czujnik_natezenia_światła"
   TextField "Text field_20" at 549,313 size 86x22; Text 'AKTUALNA / AKTUALNE'
   TextField "Text field_23" at 616,150 size 32x18; Text '2'
   TextField "Text field_24" at 614,205 size 32x18; Text '2'
   Bar "Bar_5" at 656,111 size 45x250; MinimumValue 400; MaximumValue 950
      ProcessValue <- "Poziom_CO2_auto"
   TextField "Text field_21" at 656,65 size 128x23; Text 'SYSTEM OKIEN / POZIOM CO2'
   IOField "I/O field_9" at 723,254 size 66x40; FormatPattern 999
      ProcessValue <- "Poziom_CO2_auto"
   TextField "Text field_22" at 699,216 size 101x22; Text 'USTAWIONA / USTAWIONE'
   IOField "I/O field_10" at 723,333 size 62x40; FormatPattern 999
      ProcessValue <- "Wewnetrzny_czujnik_CO2"
   TextField "Text field_25" at 708,314 size 86x22; Text 'AKTUALNA'
   Button "Button_6" at 714,134 size 73x40; TextOff '+ / +25ppm'
      on Click: function_dd21b452("Poziom_CO2_auto", 25)
   Button "Button_12" at 714,186 size 73x40; TextOff '+ / -25ppm'
      on Click: function_b9b71300("Poziom_CO2_auto", 25)
   GraphicView "Graphic view_5" at 754,83 size 40x40; Picture "sensor_2828470"
   GraphicView "Graphic view_6" at 17,400 size 55x55; Picture "window_11250237"

screen "Symulacja_czujnikow" 800x480
   TextField "Text field_1" at 12,58 size 252x23; Text 'Czujnik Wilgotności powietrza'
   TextField "Text field_2" at 306,58 size 214x23; Text 'Czujnik Wilgotności gleby'
   TextField "Text field_3" at 32,202 size 202x23; Text 'Termometr wewnętrzny'
   TextField "Text field_4" at 323,202 size 197x23; Text 'Termometr zewnętrzny'
   TextField "Text field_5" at 566,58 size 216x23; Text 'Czujnik natężenia światła'
   TextField "Text field_6" at 607,202 size 124x23; Text 'Czujnik wiatru'
   TextField "Text field_7" at 27,346 size 208x23; Text 'Wewnętrzny czujnik CO2'
   TextField "Text field_8" at 306,346 size 202x23; Text 'Zewnętrzny czujnik CO2'
   TextField "Text field_9" at 569,346 size 206x23; Text 'Stopień zasłonięcia rolet'
   IOField "I/O field_4" at 599,94 size 150x60; FormatPattern 9999
      ProcessValue <- "Czujnik_natezenia_światła"
   IOField "I/O field_5" at 599,242 size 150x60; FormatPattern 999
      ProcessValue <- "Czujnik_wiatru"
   IOField "I/O field_6" at 69,375 size 150x60; FormatPattern 9999
      ProcessValue <- "Wewnetrzny_czujnik_CO2"
   IOField "I/O field_7" at 346,375 size 150x60; FormatPattern 9999
      ProcessValue <- "Zewnetrzny_czujnik_CO2"
   IOField "I/O field_8" at 599,375 size 150x60; FormatPattern 999
      ProcessValue <- "Stopien_zasloniecia_rolet"
   IOField "I/O field_10" at 69,94 size 150x60; FormatPattern 999
      ProcessValue <- "Czujnik_wilgotności_powietrza"
   IOField "I/O field_11" at 346,94 size 150x60; FormatPattern 999
      ProcessValue <- "Czujnik_wilgotności_gleby"
   IOField "I/O field_12" at 69,242 size 150x60; FormatPattern 99.9
      ProcessValue <- "Temperatura_wewnetrzna"
   IOField "I/O field_13" at 346,242 size 150x60; FormatPattern 99.9
      ProcessValue <- "Temperatura_zewnetrzna"
   TextField "Text field_10" at 248,5 size 321x34; Text 'ZAPISZ RECEPTURE / SYMULACJA CZUJNIKÓW'
   Button "Button_1" at 750,0 size 50x50; TextOff 'WRÓĆ'; PictureOff "Back_arrow"
      on Click: function_efd93a16()
   Button "Button_14" at 3,1 size 43x43; TextOff 'DOM'; PictureOff "home_1"
      on Click: ActivateScreen("Root screen", 0)

screen "Root screen" 800x480, template "Template_1"
   on GenerateScreen: SetTag("Tag_ScreenNumber", 0)
   Button "Button_1" at 9,154 size 300x70; TextOff 'TRYB MANUALNY'
      on Click: ActivateScreen("tryb_manualny", 0)
   Button "Button_2" at 10,70 size 300x70; TextOff 'TRYB AUTOMATYCZNY'
      on Click: ActivateScreen("tryb_automatyczny", 0)
   TextField "Text field_2" at 73,1 size 601x52; Text 'AUTOMATYCZNA SZKLARNIA'
   GraphicView "Graphic view_1" at 370,70 size 392x338; Picture "garden-tools-graphic-clipart-design-free-png"
   Button "Button_5" at 10,237 size 300x70; TextOff 'TRYB RECEPTUR'
      on Click: function_e3503463('\USB_X60.1\record.csv', U 0, 2, 1, N); ActivateScreen("Receptury", 0)
   Button "Button_3" at 10,322 size 300x70; TextOff 'SYMULACJA'
      on Click: ActivateScreen("Symulacja_czujnikow", 0)

